HMI tags "Tabla de variables estándar_1"
   "MC066_STD" : , 1 s
   "MV031_STD" : , 1 s
   "MV032_STD" : , 1 s
   "MV030_STD" : , 1 s
   "DIP_1" : , internal
   "MP016_STD" : , 1 s
   "MC004_STD" : , 1 s
   "MP013_STD" : , 1 s
   "MV033_STD" : , 1 s
   "MC001_STD" : , 1 s
   "MC060_STD" : , 1 s
   "MC002_STD" : , 1 s
   "MP012_STD" : , 1 s
   "MC065_STD" : , 1 s
   "MS051_STD" : , 1 s
   "MC006_STD" : , 1 s
   "MP011_STD" : , 1 s
   "Iluminati_STD" : , 1 s
   "MC064_STD" : , 1 s
   "MS052_STD" : , 1 s
   "MT010_STD" : , 1 s
   "MS053_STD" : , 1 s
   "MP019_STD" : , 1 s
   "MC005_STD" : , 1 s
   "MC061_STD" : , 1 s
   "MV034_STD" : , 1 s
   "MC063_STD" : , 1 s
   "MP015_STD" : , 1 s
   "MT007_STD" : , 1 s
   "MS055_STD" : , 1 s
   "MP018_STD" : , 1 s
   "MP014_STD" : , 1 s
   "MS054_STD" : , 1 s
   "MS050_STD" : , 1 s
   "MP010_STD" : , 1 s
   "MT008_STD" : , 1 s
   "MT009_STD" : , 1 s
   "MC003_STD" : , 1 s
   "MC062_STD" : , 1 s
   "EB5" : Word, 1 s
   "EB7" : Word, 1 s
   "EB4" : Word, 1 s
   "EW8" : Word, 1 s
   "ACK_ALARMA_2" : Int, 1 s
   "MP020_STD" : Word, 1 s
   "MP021_STD" : Word, 1 s
   "MP022_STD" : Word, 1 s
   "CERO" : Bool, 1 s
   "UNO" : Bool, 1 s
   "IndCh" : Bool, 1 s
   "IndTrCh" : Bool, 1 s
   "IndCmpBaja" : Bool, 1 s
   "IndSecBaja" : Bool, 1 s
   "IndCmpAlta" : Bool, 1 s
   "IndSecAlta" : Bool, 1 s
   "IndTrCav" : Bool, 1 s
   "AnularSirena?" : Bool, internal
   "HorasBoost1" : DInt, 1 s
   "HorasBoost2" : DInt, 1 s
   "BoostPrHoras" : Bool, 1 s
   "BoostInvP" : Bool, 1 s
   "PrioridadBoost1" : Int, 1 s
   "PrioridadBoost2" : Int, 1 s
   "BoostInvPMan" : Bool, 1 s
   "min_boost1" : Int, 1 s
   "SegsBoost1" : Int, 1 s
   "SegsBoost" : Int, 1 s
   "MinBoost2" : Int, 1 s
   "FT1_AGUA" : Bool = PLC "FT1_AGUA", 1 s

HMI tags "AlarmasMTA"
   "AlarmasWord0" : Int, 1 s
   "AlarmasWord1" : Int, 1 s
   "AlarmasWord2" : Int, 1 s
   "AlarmasWord3" : Int, 1 s
   "AlarmasWord4" : Int, 1 s
   "AlarmasWord5" : Int, 1 s
   "AlarmasWord6" : Int, 1 s
   "AlarmasWord7" : Int, 1 s
   "AlarmasWord8" : Int, 1 s
   "Rec0" : Int, 1 s
   "Rec1" : Int, 1 s
   "Rec2" : Int, 1 s
   "Rec3" : Int, 1 s
   "Rec4" : Int, 1 s
   "Rec5" : Int, 1 s
   "Rec6" : Int, 1 s
   "Rec7" : Int, 1 s
   "Rec8" : Int, 1 s
   "AlarmasWord9" : Int, 1 s
   "AlarmasWord10" : Int, 1 s
   "AlarmasWord11" : Int, 1 s
   "AlarmasWord12" : Int, 1 s
   "AlarmasWord13" : Int, 1 s
   "AlarmasWord14" : Int, 1 s
   "Rec9" : Int, 1 s
   "Rec10" : Int, 1 s
   "Rec11" : Int, 1 s
   "Rec12" : Int, 1 s
   "Rec13" : Int, 1 s
   "Rec14" : Int, 1 s
   "AlarmasWord15" : Int, 1 s
   "Rec15" : Int, 1 s
   "ReconocerTODAS" : Bool, 1 s
   "EncendidoPLC" : Bool, 1 s
   "AlarmasWord16" : Int, 1 s
   "Rec16" : Int, 1 s
   "ReconocerTODAS_1" : Bool, 1 s
   "AlarmasWord18" : Int, 1 s
   "Rec18" : Int, 1 s
   "AlarmasWord19" : Int, 1 s
   "Rec19" : Int, 1 s
   "AlarmasWord20" : Int, 1 s
   "AlarmasWord21" : Int, 1 s
   "AlarmasWord22" : Int, 1 s
   "AlarmasWord23" : Int, 1 s
   "AlarmasWord24" : Int, 1 s
   "Rec20" : Int, 1 s
   "Rec21" : Int, 1 s
   "Rec22" : Int, 1 s
   "Rec23" : Int, 1 s
   "Rec24" : Int, 1 s

HMI tags "AutoTorresCav"
   "AutoV030" : Bool, 1 s
   "AutoV031" : Bool, 1 s
   "SP-OFF-V030" : Int, 1 s
   "SP-OFF-V031" : Int, 1 s
   "SP-ON-V030" : Int, 1 s
   "SP-ON-V031" : Int, 1 s

HMI tags "AutoTorresChillers"
   "AutoV001" : Bool, 1 s
   "AutoV002" : Bool, 1 s
   "AutoV003" : Bool, 1 s
   "SP-ON-V001" : Int, 1 s
   "SP-ON-V002" : Int, 1 s
   "SP-ON-V003" : Int, 1 s
   "SP-OFF-V001" : Int, 1 s
   "SP-OFF-V002" : Int, 1 s
   "SP-OFF-V003" : Int, 1 s
   "TemperaturatorresCH" : Real, 1 s

HMI tags "Booster"
   "AlarmaBooster" : Bool, 1 s
   "Booster_ModoManten" : Bool, 1 s
   "Booster_ModoManual" : Bool, 1 s
   "Booster_ModoAutoma" : Bool, 1 s
   "Booster_PlsManten" : Bool, 1 s
   "Booster_PlsManual" : Bool, 1 s
   "Booster_PlsAutoma" : Bool, 1 s
   "AnimaMotBooster" : Byte, 1 s
   "BoosterOrdMarcha" : Bool, 1 s
   "Booster_Conf_Marcha" : Bool, 1 s
   "Booster_Presost_Ctrl" : Bool, 1 s
   "Booster_Presost_PA" : Bool, 1 s
   "Booster_Habilitacion" : Bool, 1 s
   "Booster2_Conf_Marcha" : Bool, 1 s
   "Booster2_Habilitacion" : Bool, 1 s
   "Booster2_ModoAutoma" : Bool, 1 s
   "Booster2_ModoManten" : Bool, 1 s
   "Booster2_ModoManual" : Bool, 1 s
   "Booster2_PlsAutoma" : Bool, 1 s
   "Booster2_PlsManten" : Bool, 1 s
   "Booster2_PlsManual" : Bool, 1 s
   "AnimaMotBooster2" : Byte, 1 s
   "Booster2OrdMarcha" : Bool, 1 s
   "TiempoAyudaON" : Int, 1 s
   "TiempoAyudaOFF" : Int, 1 s
   "DifHorINVBoost" : DInt, 1 s
   "LimArrBoostPrio2" : Real, 1 s
   "LimArrBoostPrio1" : Real, 1 s
   "LimParBoostPrio2" : Real, 1 s
   "LimParBoostPrio1" : Real, 1 s
   "Presión_Actual_Boosters" : Real, 1 s
   "Ctrl_Analógico" : Bool, 1 s
   "Ver_Config" : Bool, internal
   "CotaSupPresAna" : Real, 1 s

HMI tags "CFG-Analog-MTA"
   "PresiónALTA" : Real, 1 s
   "PresiónBAJA" : Real, 1 s
   "TempCAV" : Real, 1 s
   "TempCH" : Real, 1 s
   "CFG-ALtaHH" : Real, 1 s
   "CFG-ALtaH" : Real, 1 s
   "CFG-ALtaL" : Real, 1 s
   "CFG-ALtaLL" : Real, 1 s
   "CFG-BajaHH" : Real, 1 s
   "CFG-BajaH" : Real, 1 s
   "CFG-BajaL" : Real, 1 s
   "CFG-BajaLL" : Real, 1 s
   "LO_potencia" : Real, 1 s
   "HI_caudal" : Real, 1 s
   "LO_caudal" : Real, 1 s
   "HI_potencia" : Real, 1 s
   "Caudal" : Real, 1 s
   "Potencia" : Real, 1 s

HMI tags "ChillersMTA"
   "HabMT007" : Bool, 1 s
   "HabMT008" : Bool, 1 s
   "HabMT009" : Bool, 1 s
   "HabMT010" : Bool, 1 s
   "DesMT007" : Bool, 1 s
   "DesMT008" : Bool, 1 s
   "DesMT009" : Bool, 1 s
   "DesMT010" : Bool, 1 s
   "MarchaMT007" : Bool, 1 s
   "MarchaMT008" : Bool, 1 s
   "MarchaMT009" : Bool, 1 s
   "MarchaMT010" : Bool, 1 s
   "ParadaMT007" : Bool, 1 s
   "ParadaMT008" : Bool, 1 s
   "ParadaMT009" : Bool, 1 s
   "ParadaMT010" : Bool, 1 s
   "Habilitación-CH-SOP-GR" : Bool, 1 s
   "Habilitación-CH-SOP-CH" : Bool, 1 s
   "Habilitación-CH-ENV-GR" : Bool, 1 s
   "Habilitación-CH-ENV-CH" : Bool, 1 s
   "Alarma1-CH-SOP-GR" : Bool, 1 s
   "Alarma2-CH-SOP-GR" : Bool, 1 s
   "RUN-CH-SOP-GR" : Bool, 1 s
   "MAX-CH-SOP-GR" : Bool, 1 s
   "AnimaciónMT007" : Byte, 1 s
   "AnimaciónMT008" : Byte, 1 s
   "AnimaciónMT009" : Byte, 1 s
   "AnimaciónMT010" : Byte, 1 s
   "AnimaciónMP010" : Byte, 1 s
   "AnimaciónMP011" : Byte, 1 s
   "AnimaciónMP012" : Byte, 1 s
   "AnimaciónMP013" : Byte, 1 s
   "HabMP010" : Bool, 1 s
   "HabMP011" : Bool, 1 s
   "HabMP012" : Bool, 1 s
   "HabMP013" : Bool, 1 s
   "HabMP018" : Bool, 1 s
   "HabMP019" : Bool, 1 s
   "DesMP010" : Bool, 1 s
   "DesMP011" : Bool, 1 s
   "DesMP012" : Bool, 1 s
   "DesMP013" : Bool, 1 s
   "DesMP018" : Bool, 1 s
   "DesMP019" : Bool, 1 s
   "MarchaMP010" : Bool, 1 s
   "MarchaMP011" : Bool, 1 s
   "MarchaMP012" : Bool, 1 s
   "MarchaMP013" : Bool, 1 s
   "MarchaMP018" : Bool, 1 s
   "MarchaMP019" : Bool, 1 s
   "ParadaMP010" : Bool, 1 s
   "ParadaMP011" : Bool, 1 s
   "ParadaMP012" : Bool, 1 s
   "ParadaMP013" : Bool, 1 s
   "ParadaMP018" : Bool, 1 s
   "ParadaMP019" : Bool, 1 s
   "AnimaciónMP018" : Byte, 1 s
   "AnimaciónMP019" : Byte, 1 s
   "DesV001" : Bool, 1 s
   "DesV002" : Bool, 1 s
   "HabV001" : Bool, 1 s
   "HabV002" : Bool, 1 s
   "MarchaV001" : Bool, 1 s
   "MarchaV002" : Bool, 1 s
   "ParadaV001" : Bool, 1 s
   "ParadaV002" : Bool, 1 s
   "AnimaciónV001" : Byte, 1 s
   "AnimaciónV002" : Byte, 1 s
   "VentiladoresMTA" : Bool, internal
   "MAX-CH-ENV-GR" : Bool, 1 s
   "RUN-CH-ENV-GR" : Bool, 1 s
   "Alarma2-CH-ENV-GR" : Bool, 1 s
   "Alarma1-CH-ENV-GR" : Bool, 1 s
   "SirenaM1" : Bool, 1 s
   "SirenaM2" : Bool, 1 s
   "SirenaM3" : Bool, 1 s
   "SirenaM4" : Bool, 1 s
   "AnimaciónV003" : Byte, 1 s
   "HabV003" : Bool, 1 s
   "DesV003" : Bool, 1 s
   "MarchaV003" : Bool, 1 s
   "ParadaV003" : Bool, 1 s
   "BombaTorreON" : Bool, 1 s
   "SirenaM5" : Bool, 1 s
   "SirenaChillers" : Bool, 1 s
   "SirenaM6" : Bool, 1 s
   "SirenaM7" : Bool, 1 s
   "SirenaM8" : Bool, 1 s
   "SirenaM9" : Bool, 1 s
   "SirenaM10" : Bool, 1 s
   "AlarmaNueva" : Bool, 1 s
   "AlarmaPresente" : Bool, 1 s
   "SinAlarmas" : Bool, 1 s
   "AlarmaAceite-CH-ENV-CH" : Bool, 1 s
   "AlarmaTemp-CH-ENV-CH" : Bool, 1 s
   "RUN-CH-ENV-CH" : Bool, 1 s
   "VerCh1MTA" : Bool, internal
   "VerCh2MTA" : Bool, internal
   "VerCh3MTA" : Bool, internal
   "VerCh4MTA" : Bool, internal
   "AlarmaPRUEBA" : DWord, 1 s
   "Presosato" : Bool, 1 s
   "CH-SOP-CH-CTC1ON" : Bool, 1 s
   "CH-SOP-CH-CTC2ON" : Bool, 1 s
   "CH-SOP-CH-TERM1" : Bool, 1 s
   "CH-SOP-CH-TERM2" : Bool, 1 s
   "CH-ENV-CH-ACT" : Bool, 1 s
   "CH-ENV-CH-TEMP" : Bool, 1 s
   "CH-ENV-CH-TERM" : Bool, 1 s
   "CH-ENV-CH-RUN" : Bool, 1 s
   "BombaTorreON2" : Bool, 1 s
   "HabV001(1)" : Bool, 1 s
   "HabV002(1)" : Bool, 1 s
   "HabV003(1)" : Bool, 1 s
   "HabV4" : Bool, 1 s
   "MarchaV001(1)" : Bool, 1 s
   "MarchaV002(1)" : Bool, 1 s
   "MarchaV003(1)" : Bool, 1 s
   "ParadaV001(1)" : Bool, 1 s
   "ParadaV002(1)" : Bool, 1 s
   "ParadaV003(1)" : Bool, 1 s
   "AnimaMenuV001" : Int, 1 s
   "AnimaMenuV002" : Int, 1 s
   "AnimaMenuV003" : Int, 1 s
   "DeshV001" : Bool, 1 s
   "DeshV002" : Bool, 1 s
   "DeshV003" : Bool, 1 s

HMI tags "CompBajaMTA"
   "HabilitaciónMC060" : Bool, 1 s
   "HabilitaciónMC061" : Bool, 1 s
   "HabilitaciónMC062" : Bool, 1 s
   "HabilitaciónMC063" : Bool, 1 s
   "HabilitaciónMC064" : Bool, 1 s
   "HabilitaciónMC065" : Bool, 1 s
   "DeshabilitaciónMC060" : Bool, 1 s
   "DeshabilitaciónMC061" : Bool, 1 s
   "DeshabilitaciónMC062" : Bool, 1 s
   "DeshabilitaciónMC063" : Bool, 1 s
   "DeshabilitaciónMC064" : Bool, 1 s
   "DeshabilitaciónMC065" : Bool, 1 s
   "MarchaMC060" : Bool, 1 s
   "MarchaMC061" : Bool, 1 s
   "MarchaMC062" : Bool, 1 s
   "MarchaMC063" : Bool, 1 s
   "MarchaMC064" : Bool, 1 s
   "MarchaMC065" : Bool, 1 s
   "ParadaMC060" : Bool, 1 s
   "ParadaMC061" : Bool, 1 s
   "ParadaMC062" : Bool, 1 s
   "ParadaMC063" : Bool, 1 s
   "ParadaMC064" : Bool, 1 s
   "ParadaMC065" : Bool, 1 s
   "AnimaMC060" : Byte, 1 s
   "AnimaMC061" : Byte, 1 s
   "AnimaMC062" : Byte, 1 s
   "AnimaMC063" : Byte, 1 s
   "AnimaMC064" : Byte, 1 s
   "AnimaMC065" : Byte, 1 s
   "VerMC060" : Bool, internal
   "VerMC061" : Bool, internal
   "VerMC062" : Bool, internal
   "VerMC063" : Bool, internal
   "VerMC064" : Bool, internal
   "MantM060" : Bool, 1 s
   "MantM061" : Bool, 1 s
   "MantM062" : Bool, 1 s
   "MantM063" : Bool, 1 s
   "MantM064" : Bool, 1 s
   "AutoMC060" : Bool, 1 s
   "AutoMC061" : Bool, 1 s
   "AutoMC062" : Bool, 1 s
   "AutoMC063" : Bool, 1 s
   "AutoMC064" : Bool, 1 s
   "SponMC060" : Real, 1 s
   "SponMC061" : Real, 1 s
   "SponMC062" : Real, 1 s
   "SponMC063" : Real, 1 s
   "SponMC064" : Real, 1 s
   "SpoffMC060" : Real, 1 s
   "SpoffMC061" : Real, 1 s
   "SpoffMC062" : Real, 1 s
   "SpoffMC063" : Real, 1 s
   "SpoffMC064" : Real, 1 s
   "AnimMenuMC060" : Int, 1 s
   "AnimMenuMC061" : Int, 1 s
   "AnimMenuMC062" : Int, 1 s
   "AnimMenuMC063" : Int, 1 s
   "AnimMenuMC064" : Int, 1 s
   "HabilitarMC060" : Bool, 1 s
   "AnularSirenaCav" : Bool, 1 s
   "VerMC65" : Bool, internal

HMI tags "CompresoresAltaMTA"
   "Sop1" : Bool, 1 s
   "Sop2" : Bool, 1 s
   "Sop3" : Bool, 1 s
   "ReqSop1" : Int, 1 s
   "ReqSop2" : Int, 1 s
   "ReqSop3" : Int, 1 s
   "NinSop" : Bool, 1 s
   "VCMP1" : Int, 1 s
   "VCMP2" : Int, 1 s
   "VCMP3" : Int, 1 s
   "VCMP4" : Int, 1 s
   "VCMP5" : Int, 1 s
   "IncP1" : Bool, 100 ms
   "IncP2" : Bool, 100 ms
   "IncP3" : Bool, 100 ms
   "IncP4" : Bool, 100 ms
   "IncP5" : Bool, 100 ms
   "DecP1" : Bool, 1 s
   "DecP2" : Bool, 1 s
   "DecP3" : Bool, 1 s
   "DecP4" : Bool, 1 s
   "DecP5" : Bool, 1 s
   "PriRealCMP1" : Int, 1 s
   "PriRealCMP2" : Int, 1 s
   "PriRealCMP3" : Int, 1 s
   "PriRealCMP4" : Int, 1 s
   "PriRealCMP5" : Int, 1 s
   "Auto1" : Bool, 1 s
   "Auto2" : Bool, 1 s
   "Auto3" : Bool, 1 s
   "Auto4" : Bool, 1 s
   "Auto5" : Bool, 1 s
   "IndV1" : Bool, 100 ms
   "IndV2" : Bool, 100 ms
   "IndV3" : Bool, 100 ms
   "IndV4" : Bool, 100 ms
   "IndV5" : Bool, 100 ms
   "IndR1" : Bool, 100 ms
   "IndR2" : Bool, 100 ms
   "IndR3" : Bool, 100 ms
   "IndR4" : Bool, 100 ms
   "IndR5" : Bool, 100 ms
   "Est1" : Word, 1 s
   "Est2" : Word, 1 s
   "Est3" : Word, 1 s
   "Est4" : Word, 1 s
   "Est5" : Word, 1 s
   "LimSUP1" : Real, 1 s
   "LimSUP2" : Real, 1 s
   "LimSUP3" : Real, 1 s
   "LimSUP4" : Real, 1 s
   "LimSUP5" : Real, 1 s
   "LimINF1" : Real, 1 s
   "LimINF2" : Real, 1 s
   "LimINF3" : Real, 1 s
   "LimINF4" : Real, 1 s
   "LimINF5" : Real, 1 s
   "PresMaX" : Real, 1 s
   "Delta" : Real, 1 s
   "Hist" : Real, 1 s
   "CompReq" : Int, 1 s
   "CompReqINI" : Int, 1 s
   "AnimMenuMC001" : Int, 1 s
   "AnimMenuMC002" : Int, 1 s
   "AnimMenuMC003" : Int, 1 s
   "AnimMenuMC004" : Int, 1 s
   "AnimMenuMC005" : Int, 1 s
   "SPON1" : Real, 1 s
   "SPON2" : Real, 1 s
   "SPON3" : Real, 1 s
   "SPON4" : Real, 1 s
   "SPON5" : Real, 1 s
   "SPOFF1" : Real, 1 s
   "SPOFF2" : Real, 1 s
   "SPOFF3" : Real, 1 s
   "SPOFF4" : Real, 1 s
   "SPOFF5" : Real, 1 s
   "MantMC001" : Bool, 1 s
   "MantMC002" : Bool, 1 s
   "MantMC003" : Bool, 1 s
   "MantMC004" : Bool, 1 s
   "MantMC005" : Bool, 1 s
   "IndVparp1" : Bool, 1 s
   "IndVparp2" : Bool, 1 s
   "IndVparp3" : Bool, 1 s
   "IndVparp4" : Bool, 1 s
   "IndVparp5" : Bool, 1 s
   "TiempoenVacío" : Int, 1 s
   "TiemposinReq" : Int, 1 s
   "TiempoSop" : Int, 1 s
   "HistCRT" : Real, 1 s
   "LimINFCRT" : Real, 1 s
   "LimSUPCRT" : Real, 1 s
   "PanMCH1" : Bool, 1 s
   "PanMCH2" : Bool, 1 s
   "PanMCH3" : Bool, 1 s
   "PanMCH4" : Bool, 1 s
   "PanMCH5" : Bool, 1 s
   "MarchaMC001" : Bool, 1 s
   "MarchaMC002" : Bool, 1 s
   "MarchaMC003" : Bool, 1 s
   "MarchaMC004" : Bool, 1 s
   "MarchaMC005" : Bool, 1 s
   "ParadaMC001" : Bool, 1 s
   "ParadaMC002" : Bool, 1 s
   "ParadaMC003" : Bool, 1 s
   "ParadaMC004" : Bool, 1 s
   "ParadaMC005" : Bool, 1 s
   "AnimMotorMC001" : Byte, 1 s
   "AnimMotorMC002" : Byte, 1 s
   "AnimMotorMC003" : Byte, 1 s
   "AnimMotorMC004" : Byte, 1 s
   "AnimMotorMC005" : Byte, 1 s
   "EV1" : Bool, 1 s
   "EV2" : Bool, 1 s
   "EV3" : Bool, 1 s
   "EV4" : Bool, 1 s
   "EV5" : Bool, 1 s
   "HORAS1" : DInt, 1 s
   "HORAS2" : DInt, 1 s
   "HORAS3" : DInt, 1 s
   "HORAS4" : DInt, 1 s
   "HORAS5" : DInt, 1 s
   "MIN1" : Int, 1 s
   "MIN2" : Int, 1 s
   "MIN3" : Int, 1 s
   "MIN4" : Int, 1 s
   "MIN5" : Int, 1 s
   "MarchaOK1" : Bool, 1 s
   "MarchaOK2" : Bool, 1 s
   "MarchaOK3" : Bool, 1 s
   "MarchaOK4" : Bool, 1 s
   "MarchaOK5" : Bool, 1 s
   "ForzarMarcha1" : Bool, 1 s
   "ForzarMarcha2" : Bool, 1 s
   "ForzarMarcha3" : Bool, 1 s
   "ForzarMarcha4" : Bool, 1 s
   "ForzarMarcha5" : Bool, 1 s
   "ForzarParada1" : Bool, 1 s
   "ForzarParada2" : Bool, 1 s
   "ForzarParada3" : Bool, 1 s
   "ForzarParada4" : Bool, 1 s
   "ForzarParada5" : Bool, 1 s
   "SPONF1" : Real, 1 s
   "SPONF2" : Real, 1 s
   "SPONF3" : Real, 1 s
   "SPONF4" : Real, 1 s
   "SPONF5" : Real, 1 s
   "SPOFFF1" : Real, 1 s
   "SPOFFF2" : Real, 1 s
   "SPOFFF3" : Real, 1 s
   "SPOFFF4" : Real, 1 s
   "SPOFFF5" : Real, 1 s
   "ForzandoMarcha1" : Bool, 1 s
   "ForzandoMarcha2" : Bool, 1 s
   "ForzandoMarcha3" : Bool, 1 s
   "ForzandoMarcha4" : Bool, 1 s
   "ForzandoMarcha5" : Bool, 1 s
   "MediaCargaBellis" : Bool, 1 s
   "SPONF3b" : Real, 1 s
   "SPOFFF3b" : Real, 1 s
   "EV3b" : Bool, 1 s
   "TiempoMaxBellismedia" : Int, 1 s
   "Est6" : Int, 1 s
   "PriRealCMP6" : Int, 1 s
   "IndV6" : Bool, 1 s

HMI tags "IluminaciónMTA"
   "TiempoIluminación" : Word, 1 s
   "EncendidoPanel" : Bool, 1 s
   "ApagadoPanel" : Bool, 1 s
   "ON" : Bool, 1 s
   "MantenerON" : Bool, 1 s
   "AlarmaBoosters" : Bool, 1 s

HMI tags "SecadoresAltaMTA"
   "AnimaMS050" : Byte, 1 s
   "AnimaMS051" : Byte, 1 s
   "AnimaMS052" : Byte, 1 s
   "AnimaMS053" : Byte, 1 s
   "DeshabilitaciónMS050" : Bool, 1 s
   "DeshabilitaciónMS051" : Bool, 1 s
   "DeshabilitaciónMS052" : Bool, 1 s
   "DeshabilitaciónMS053" : Bool, 1 s
   "HabilitaciónMS050" : Bool, 1 s
   "HabilitaciónMS051" : Bool, 1 s
   "HabilitaciónMS052" : Bool, 1 s
   "HabilitaciónMS053" : Bool, 1 s
   "MantMS050" : Bool, 1 s
   "MantMS051" : Bool, 1 s
   "MantMS052" : Bool, 1 s
   "MantMS053" : Bool, 1 s
   "MarchaMS050" : Bool, 1 s
   "MarchaMS051" : Bool, 1 s
   "MarchaMS052" : Bool, 1 s
   "MarchaMS053" : Bool, 1 s
   "ParadaMS050" : Bool, 1 s
   "ParadaMS051" : Bool, 1 s
   "ParadaMS052" : Bool, 1 s
   "ParadaMS053" : Bool, 1 s
   "AnimaMenuMS050" : Int, 1 s
   "AnimaMenuMS051" : Int, 1 s
   "AnimaMenuMS052" : Int, 1 s
   "AnimaMenuMS053" : Int, 1 s
   "Enc1MS050" : Int, 1 s
   "Enc2MS050" : Int, 1 s
   "Enc1MS051" : Int, 1 s
   "Enc2MS051" : Int, 1 s
   "Enc1MS052" : Int, 1 s
   "Enc2MS052" : Int, 1 s
   "Enc1MS053" : Int, 1 s
   "Enc2MS053" : Int, 1 s
   "AutoMS050" : Bool, 1 s
   "AutoMS051" : Bool, 1 s
   "AutoMS052" : Bool, 1 s
   "AutoMS053" : Bool, 1 s

HMI tags "SecadoresBaja"
   "AnimaMS054" : Byte, 1 s
   "AnimaMS055" : Byte, 1 s
   "DeshabilitaciónMS054" : Bool, 1 s
   "DeshabilitaciónMS055" : Bool, 1 s
   "HabilitaciónMS054" : Bool, 1 s
   "HabilitaciónMS055" : Bool, 1 s
   "MarchaMS054" : Bool, 1 s
   "MarchaMS055" : Bool, 1 s
   "ParadaMS054" : Bool, 1 s
   "ParadaMS055" : Bool, 1 s
   "MantMS054" : Bool, 1 s
   "MantMS055" : Bool, 1 s

HMI tags "SENTRON PAC 3200"
   "Tension Fase R" : Float, 1 s
   "Tension fase S" : Float, 1 s
   "Tension Fase T" : Float, 1 s
   "Tension Linea RS" : Float, 1 s
   "Tension Linea ST" : Float, 1 s
   "Tension Linea TR" : Float, 1 s
   "Corriente fase R" : Float, 1 s
   "Corriente Fase S" : Float, 1 s
   "Corriente Fase T" : Float, 1 s
   "Pot.Apa R" : Float, 1 s
   "Pot.Apa S" : Float, 1 s
   "Pot.Apa T" : Float, 1 s
   "Pot.Act R" : Float, 1 s
   "Pot.Act S" : Float, 1 s
   "Pot.Act T" : Float, 1 s
   "Pot.ReAct R" : Float, 1 s
   "Pot.ReAct S" : Float, 1 s
   "Pot.ReAct T" : Float, 1 s
   "Coseno R" : Float, 1 s
   "Coseno S" : Float, 1 s
   "Coseno T" : Float, 1 s
   "THD-R TensionFase R" : Float, 1 s
   "THD-R Tension Fase S" : Float, 1 s
   "THD-R Tension Fase T" : Float, 1 s
   "THD-R Corriente Fase R" : Float, 1 s
   "THD-R Corriente Fase S" : Float, 1 s
   "THD-R Corriente Fase T" : Float, 1 s
   "Frecuencia" : Float, 1 s
   "Tension Media Fase" : Float, 1 s
   "Tension Media de Linea" : Float, 1 s
   "Corriente Media" : Float, 1 s
   "Pot Apa Total" : Float, 1 s
   "Pot Act Total" : Float, 1 s
   "Pot ReAct Total" : Float, 1 s
   "coseno Total" : Float, 1 s
   "desbalance de tension" : Float, 1 s
   "desbalance de corriente" : Float, 1 s
   "Tension Maxima R" : Float, 1 s
   "Tension Maxima S" : Float, 1 s
   "Tension Maxima T" : Float, 1 s
   "Tension Maxima RS" : Float, 1 s
   "Tension Maxima ST" : Float, 1 s
   "Tension Maxima TR" : Float, 1 s
   "Corriente Maxima R" : Float, 1 s
   "Corriente Maxima S" : Float, 1 s
   "Corriente Maxima T" : Float, 1 s

HMI tags "TorresCav-MTA"
   "AnimaMV030" : Byte, 1 s
   "AnimaMV031" : Byte, 1 s
   "AnimaMP014" : Byte, 1 s
   "AnimaMP015" : Byte, 1 s
   "DeshabilitaciónMV030" : Bool, 1 s
   "DeshabilitaciónMV031" : Bool, 1 s
   "DeshabilitaciónMP014" : Bool, 1 s
   "DeshabilitaciónMP015" : Bool, 1 s
   "HabilitaciónMV030" : Bool, 1 s
   "HabilitaciónMV031" : Bool, 1 s
   "HabilitaciónMP014" : Bool, 1 s
   "HabilitaciónMP015" : Bool, 1 s
   "MantMV030" : Bool, 1 s
   "MantMV031" : Bool, 1 s
   "MantMP014" : Bool, 1 s
   "MantMP015" : Bool, 1 s
   "MarchaMV030" : Bool, 1 s
   "MarchaMV031" : Bool, 1 s
   "MarchaMP014" : Bool, 1 s
   "MarchaMP015" : Bool, 1 s
   "ParadaMV030" : Bool, 1 s
   "ParadaMV031" : Bool, 1 s
   "ParadaMP014" : Bool, 1 s
   "ParadaMP015" : Bool, 1 s
   "MenuV030" : Int, 1 s
   "MenuV031" : Int, 1 s

discrete alarms
   1: '', class MTA, trigger "AlarmasWord13" bit 9
   2: '', class MTA, trigger "AlarmasWord13" bit 10
   3: '', class MTA, trigger "AlarmasWord13" bit 11
   4: '', class MTA, trigger "AlarmasWord13" bit 12
   5: '', class MTA, trigger "AlarmasWord13" bit 13
   6: '', class MTA, trigger "AlarmasWord13" bit 14
   7: '', class MTA, trigger "AlarmasWord13" bit 15
   8: '', class MTA, trigger "AlarmasWord14" bit 8
   9: '', class MTA, trigger "AlarmasWord14" bit 9
   10: '', class MTA, trigger "AlarmasWord14" bit 10
   11: '', class MTA, trigger "AlarmasWord14" bit 11
   12: '', class MTA, trigger "AlarmasWord14" bit 12
   13: '', class MTA, trigger "AlarmasWord6" bit 8
   14: '', class MTA, trigger "AlarmasWord6" bit 9
   15: '', class MTA, trigger "AlarmasWord14" bit 13
   16: '', class MTA, trigger "AlarmasWord14" bit 14
   17: '', class MTA, trigger "AlarmasWord14" bit 15
   18: '', class MTA, trigger "AlarmasWord15" bit 8
   19: '', class MTA, trigger "AlarmasWord15" bit 9
   20: '', class MTA, trigger "AlarmasWord15" bit 10
   21: '', class MTA, trigger "AlarmasWord15" bit 11
   22: '', class MTA, trigger "AlarmasWord15" bit 12
   23: '', class MTA, trigger "AlarmasWord15" bit 13
   24: '', class MTA, trigger "AlarmasWord15" bit 14
   25: '', class MTA, trigger "AlarmasWord15" bit 15
   26: '', class MTA, trigger "AlarmasWord16" bit 8
   27: '', class MTA, trigger "AlarmasWord16" bit 9
   28: '', class MTA, trigger "AlarmasWord16" bit 10
   29: '', class MTA, trigger "AlarmasWord16" bit 11
   30: '', class MTA, trigger "AlarmasWord16" bit 12
   31: '', class MTA, trigger "AlarmasWord16" bit 13
   32: '', class MTA, trigger "AlarmasWord16" bit 14
   33: '', class MTA, trigger "AlarmasWord16" bit 15
   50: '', class MTA, trigger "AlarmasWord6" bit 10
   53: '', class MTA, trigger "AlarmasWord6" bit 11
   66: '', class MTA, trigger "AlarmasWord7" bit 8
   67: '', class MTA, trigger "AlarmasWord7" bit 9
   68: '', class MTA, trigger "AlarmasWord7" bit 10
   69: '', class MTA, trigger "AlarmasWord7" bit 11
   70: '', class MTA, trigger "AlarmasWord7" bit 12
   71: '', class MTA, trigger "AlarmasWord7" bit 13
   72: '', class MTA, trigger "AlarmasWord7" bit 14
   73: '', class MTA, trigger "AlarmasWord7" bit 15
   74: '', class MTA, trigger "AlarmasWord8" bit 8
   75: '', class MTA, trigger "AlarmasWord8" bit 9
   76: '', class MTA, trigger "AlarmasWord8" bit 10
   77: '', class MTA, trigger "AlarmasWord8" bit 11
   78: '', class MTA, trigger "AlarmasWord8" bit 12
   79: '', class MTA, trigger "AlarmasWord8" bit 13
   80: '', class MTA, trigger "AlarmasWord8" bit 14
   81: '', class MTA, trigger "AlarmasWord8" bit 15
   82: '', class MTA, trigger "AlarmasWord9" bit 8
   83: '', class MTA, trigger "AlarmasWord9" bit 9
   87: '', class MTA, trigger "AlarmasWord6" bit 12
   88: '', class MTA, trigger "AlarmasWord6" bit 13
   89: '', class MTA, trigger "AlarmasWord6" bit 14
   90: '', class MTA, trigger "AlarmasWord6" bit 15
   91: '', class MTA, trigger "AlarmasWord9" bit 10
   92: '', class MTA, trigger "AlarmasWord9" bit 11
   93: '', class MTA, trigger "AlarmasWord9" bit 12
   94: '', class MTA, trigger "AlarmasWord9" bit 13
   95: '', class MTA, trigger "AlarmasWord9" bit 14
   96: '', class MTA, trigger "AlarmasWord9" bit 15
   97: '', class MTA, trigger "AlarmasWord10" bit 8
   98: '', class MTA, trigger "AlarmasWord10" bit 9
   99: '', class MTA, trigger "AlarmasWord10" bit 10
   100: '', class MTA, trigger "AlarmasWord10" bit 11
   101: '', class MTA, trigger "AlarmasWord10" bit 12
   102: '', class MTA, trigger "AlarmasWord10" bit 13
   103: '', class MTA, trigger "AlarmasWord10" bit 14
   104: '', class MTA, trigger "AlarmasWord10" bit 15
   105: '', class MTA, trigger "AlarmasWord11" bit 8
   106: '', class MTA, trigger "AlarmasWord11" bit 9
   107: '', class MTA, trigger "AlarmasWord11" bit 10
   108: '', class MTA, trigger "AlarmasWord11" bit 11
   109: '', class MTA, trigger "AlarmasWord11" bit 12
   110: '', class MTA, trigger "AlarmasWord11" bit 13
   111: '', class MTA, trigger "AlarmasWord11" bit 14
   112: '', class MTA, trigger "AlarmasWord11" bit 15
   113: '', class MTA, trigger "AlarmasWord12" bit 8
   114: '', class MTA, trigger "AlarmasWord12" bit 9
   115: '', class MTA, trigger "AlarmasWord12" bit 10
   116: '', class MTA, trigger "AlarmasWord12" bit 11
   117: '', class MTA, trigger "AlarmasWord12" bit 12
   118: '', class MTA, trigger "AlarmasWord12" bit 13
   119: '', class MTA, trigger "AlarmasWord12" bit 14
   120: '', class MTA, trigger "AlarmasWord12" bit 15
   121: '', class MTA, trigger "AlarmasWord13" bit 8
   125: '', class MTA, trigger "AlarmasWord4" bit 8
   126: '', class MTA, trigger "AlarmasWord3" bit 15
   127: '', class MTA, trigger "AlarmasWord4" bit 11
   128: '', class MTA, trigger "AlarmasWord4" bit 10
   129: '', class MTA, trigger "AlarmasWord4" bit 9
   130: '', class MTA, trigger "AlarmasWord3" bit 11
   131: '', class MTA, trigger "AlarmasWord3" bit 10
   132: '', class MTA, trigger "AlarmasWord3" bit 9
   133: '', class MTA, trigger "AlarmasWord3" bit 14
   134: '', class MTA, trigger "AlarmasWord3" bit 13
   135: '', class MTA, trigger "AlarmasWord3" bit 12
   136: '', class MTA, trigger "AlarmasWord4" bit 12
   137: '', class MTA, trigger "AlarmasWord4" bit 15
   138: '', class MTA, trigger "AlarmasWord4" bit 14
   139: '', class MTA, trigger "AlarmasWord4" bit 13
   140: '', class MTA, trigger "AlarmasWord3" bit 8
   141: '', class MTA, trigger "AlarmasWord1" bit 8
   142: '', class MTA, trigger "AlarmasWord0" bit 15
   143: '', class MTA, trigger "AlarmasWord0" bit 14
   144: '', class MTA, trigger "AlarmasWord1" bit 11
   145: '', class MTA, trigger "AlarmasWord1" bit 10
   146: '', class MTA, trigger "AlarmasWord1" bit 9
   147: '', class MTA, trigger "AlarmasWord0" bit 10
   148: '', class MTA, trigger "AlarmasWord0" bit 9
   149: '', class MTA, trigger "AlarmasWord0" bit 8
   150: '', class MTA, trigger "AlarmasWord0" bit 13
   151: '', class MTA, trigger "AlarmasWord0" bit 12
   152: '', class MTA, trigger "AlarmasWord0" bit 11
   153: '', class MTA, trigger "AlarmasWord1" bit 12
   154: '', class MTA, trigger "AlarmasWord2" bit 12
   155: '', class MTA, trigger "AlarmasWord2" bit 11
   156: '', class MTA, trigger "AlarmasWord2" bit 10
   157: '', class MTA, trigger "AlarmasWord2" bit 15
   158: '', class MTA, trigger "AlarmasWord2" bit 14
   159: '', class MTA, trigger "AlarmasWord2" bit 13
   160: '', class MTA, trigger "AlarmasWord1" bit 15
   161: '', class MTA, trigger "AlarmasWord1" bit 14
   162: '', class MTA, trigger "AlarmasWord1" bit 13
   163: '', class MTA, trigger "AlarmasWord2" bit 9
   164: '', class MTA, trigger "AlarmasWord2" bit 8
   165: '', class MTA, trigger "AlarmasWord5" bit 8
   166: '', class MTA, trigger "AlarmasWord5" bit 9
   167: '', class MTA, trigger "AlarmasWord5" bit 10
   168: '', class MTA, trigger "AlarmasWord5" bit 11
   169: '', class MTA, trigger "AlarmasWord5" bit 12
   170: '', class MTA, trigger "AlarmasWord5" bit 13
   171: '', class MTA, trigger "AlarmasWord5" bit 14
   172: '', class MTA, trigger "AlarmasWord5" bit 15
   34: '', class MTA, trigger "AlarmasWord18" bit 8
   35: '', class MTA, trigger "AlarmasWord18" bit 9
   36: '', class MTA, trigger "AlarmasWord18" bit 10
   37: '', class MTA, trigger "AlarmasWord18" bit 11
   38: '', class MTA, trigger "AlarmasWord18" bit 12
   39: '', class MTA, trigger "AlarmasWord18" bit 13
   40: '', class MTA, trigger "AlarmasWord18" bit 14
   41: '', class MTA, trigger "Rec4" bit 15
   42: '', class MTA, trigger "AlarmasWord19" bit 8
   43: '', class MTA, trigger "AlarmasWord19" bit 9
   44: '', class MTA, trigger "AlarmasWord19" bit 10
   45: '', class MTA, trigger "AlarmasWord19" bit 11
   46: '', class MTA, trigger "AlarmasWord19" bit 12
   47: '', class MTA, trigger "AlarmasWord19" bit 13
   48: '', class MTA, trigger "AlarmasWord20" bit 8
   49: '', class MTA, trigger "AlarmasWord20" bit 9
   51: '', class MTA, trigger "AlarmasWord20" bit 10
   52: '', class MTA, trigger "AlarmasWord20" bit 11
   54: '', class MTA, trigger "AlarmasWord20" bit 12
   55: '', class MTA, trigger "AlarmasWord20" bit 13
   56: '', class MTA, trigger "AlarmasWord20" bit 14
   57: '', class MTA, trigger "AlarmasWord20" bit 15
   58: '', class MTA, trigger "AlarmasWord21" bit 8
   59: '', class MTA, trigger "AlarmasWord21" bit 9
   60: '', class MTA, trigger "AlarmasWord21" bit 10
   61: '', class MTA, trigger "AlarmasWord21" bit 11
   62: '', class MTA, trigger "AlarmasWord21" bit 12
   63: '', class MTA, trigger "AlarmasWord21" bit 13
   64: '', class MTA, trigger "AlarmasWord21" bit 14
   65: '', class MTA, trigger "AlarmasWord21" bit 15
   84: '', class MTA, trigger "AlarmasWord22" bit 8
   85: '', class MTA, trigger "AlarmasWord22" bit 9
   86: '', class MTA, trigger "AlarmasWord22" bit 10
   122: '', class MTA, trigger "AlarmasWord22" bit 11
   123: '', class MTA, trigger "AlarmasWord22" bit 12
   124: '', class MTA, trigger "AlarmasWord22" bit 13
   173: '', class MTA, trigger "AlarmasWord22" bit 14
   174: '', class MTA, trigger "AlarmasWord22" bit 15
   175: '', class MTA, trigger "AlarmasWord23" bit 8
   176: '', class MTA, trigger "AlarmasWord23" bit 9
   177: '', class MTA, trigger "AlarmasWord23" bit 10
   178: '', class MTA, trigger "AlarmasWord23" bit 11
   179: '', class MTA, trigger "AlarmasWord23" bit 12
   180: '', class MTA, trigger "AlarmasWord23" bit 13
   181: '', class MTA, trigger "AlarmasWord23" bit 14
   182: '', class MTA, trigger "AlarmasWord23" bit 15
   183: '', class MTA, trigger "AlarmasWord24" bit 8
   184: '', class MTA, trigger "AlarmasWord24" bit 9
   185: '', class MTA, trigger "AlarmasWord24" bit 10
   186: '', class MTA, trigger "AlarmasWord24" bit 11
   199: '', class MTA, trigger "AlarmasWord24" bit 15

text list "EstadoMotor": 0 ''; 1 ''; 2 ''; 3 ''; 4 ''; 5 ''; 6 ''; 7 ''

text list "EstadoCmpAlta": 256 ''; 512 ''; 1024 ''; 2048 ''; 4096 ''; 8192 ''; 16384 ''; 32768 ''; 1 ''

text list "Presostato Ctrl": 0 ''; 1 ''

text list "Presostato de Alarma": 0 ''; 1 ''

text list "Lista de rutas": 0 ''; 1 ''; 2 ''; 3 ''; 4 ''; 5 ''; 6 ''; 7 ''; 8 ''; 9 ''; 10 ''

text list "Lista de compresores": 0 ''; 1 ''; 2 ''; 3 ''; 4 ''; 5 ''; 6 ''; 7 ''; 8 ''; 9 ''; 10 ''

graphic list "Motor2": 0 'Motor2Dorado'; 1 'Motor2Verde_1'; 2 'Motor2VerdeOscuro'; 3 'Motor2Azul'; 4 'Motor2Celeste'; 5 'Motor2Amarillo'; 6 'Motor2Gris_1'; 7 'Motor2Rojo'; 8 'Motor2Dorado'

graphic list "MotorBelliss": 0 'dorado'; 1 'bell1ve'; 2 'bell1ve'; 3 'az'; 4 'az'; 5 'bell1am'; 6 'dorado'; 7 'az'

graphic list "BarraPrioridades": 1 'R1'; 2 'R2'; 3 'R3'; 4 'R4'; 5 'R5'; 6 'R4'; 6 'R6.rlu'

graphic list "Indicador": 0 'indDorado'; 1 'indVerde'; 2 'indVerde_1'; 3 'indAZUL'; 4 'indCeleste'; 5 'indAmarillo'; 6 'indGris'; 7 'indRojo'; 8 'indCeleste'

graphic list "BarraPrioridades_1": 1 'set1'; 2 'set2'; 3 'set3'; 4 'set4'; 5 'set5'; 6 'set4'; 6 'set6'

graphic list "BaseSullChico": 0 'BaseSullChicoDorado_4'; 1 'BaseSullChico'; 2 'BaseSullChico'; 3 'BaseSullChicoAzul_4'; 4 'BaseSullChicoAzul_4'; 5 'BaseSullChicoAmarillo_4'; 6 'BaseSullChicoGris_4'; 7 'BaseSullChicoRojo_4'; 8 'BaseSullChicoAzul_4'

graphic list "MotorTorre": 0 'torreFINAL4C2_1'; 1 'torreFINAL4C2v_2'; 2 'torreFINAL4C2v_2'; 3 'torreFINAL4C2b'; 4 'torreFINAL4C2b'; 5 'torreFINAL4C2a_2'; 6 'torreFINAL4C2_1'; 7 'torreFINAL4C2_1'

graphic list "Secador2": 0 'BaseSullChicoDorado_2'; 1 'BaseSullChico_5'; 2 'BaseSullChico_5'; 3 'BaseSullChicoAzul_2'; 4 'BaseSullChicoAzul_2'; 5 'BaseSullChicoAmarillo_2'; 6 'BaseSullChicoGris_2'; 7 'BaseSullChicoRojo_2'

graphic list "Secador1": 0 'BaseSullChicoDorado_1'; 1 'BaseSullChico_4'; 2 'BaseSullChico_4'; 3 'BaseSullChicoAzul_1'; 4 'BaseSullChicoAzul_1'; 5 'BaseSullChicoAmarillo_1'; 6 'BaseSullChicoGris_1'; 7 'BaseSullChicoRojo_1'

graphic list "Motor Grande": 0 'MotorDorado'; 1 'MotorVerde'; 2 'MotorVerde'; 3 'MotorAzul'; 4 'MotorCeleste'; 5 'MotorAmarillo'; 6 'MotorGris'; 7 'MotorRojo'; 8 'MotorCeleste'

graphic list "Mantenimiento": 0 'MECH2'; 1 'MECH1'

graphic list "Motor Chico": 0 'Booster-D-Dor2'; 1 'Booster-D-VE2'; 2 'Booster-D-VE2'; 3 'Booster-D-Azul2'; 4 'Booster-D-AZ2'; 5 'Booster-D-AM2'; 6 'Booster-D-GR'; 7 'Booster-D-RO2'; 8 'Booster-D-AZ2'

graphic list "Hélice": 0 'Booster-C1'; 1 'Booster-C2'

screen "Graf-Corrientes" 1280x800, template "Plantilla"
   TrendView "Visor de curvas_1" at 8,72 size 1260x636
   TextField "Campo de texto_16" at 493,10 size 294x27

screen "Graf-Fase" 1280x800, template "Plantilla"
   TrendView "Visor de curvas_1" at 3,65 size 1268x644
   TextField "Campo de texto_16" at 477,10 size 364x27

screen "Grafica" 1280x800, template "Plantilla"
   Button "Botón_7" at 368,280 size 240x49
   Button "Botón_12" at 367,440 size 240x49
   Button "Botón_13" at 368,216 size 240x49
   TextField "Campo de texto_1" at 55,108 size 353x27
   Button "Botón_1" at 767,280 size 240x49
   TextField "Campo de texto_16" at 521,10 size 226x27
   Button "Botón_2" at 368,344 size 240x49
   Button "Botón_3" at 766,440 size 240x49
   Button "Botón_4" at 769,526 size 240x49

screen "GraficaPALTA" 1280x800, template "Plantilla"
   TrendView "Visor de curvas_1" at 5,79 size 1234x618
   TextField "Campo de texto_16" at 521,10 size 193x27

screen "GraficaPBAJA" 1280x800, template "Plantilla"
   TrendView "Visor de curvas_1" at 5,71 size 1242x626
   TextField "Campo de texto_16" at 521,10 size 198x27

screen "GraficaTCAV" 1280x800, template "Plantilla"
   TrendView "Visor de curvas_1" at 5,71 size 1242x626
   TextField "Campo de texto_16" at 521,10 size 254x27

screen "GraficaTCH" 1280x800, template "Plantilla"
   TrendView "Visor de curvas_1" at 5,71 size 1242x626
   TextField "Campo de texto_16" at 521,10 size 243x27

screen "GraficaTodas" 1280x800, template "Plantilla"
   TrendView "Visor de curvas_1" at 5,71 size 1242x626

screen "Graf-Linea" 1280x800, template "Plantilla"
   TrendView "Visor de curvas_1" at 3,65 size 1268x652
   TextField "Campo de texto_16" at 453,10 size 370x27

screen "Graf-Pot" 1280x800, template "Plantilla"
   TrendView "Visor de curvas_1" at 3,65 size 1268x644
   TextField "Campo de texto_16" at 477,10 size 339x27

screen "Graf-PotTotal" 1280x800, template "Plantilla"
   TrendView "Visor de curvas_1" at 3,65 size 1268x644
   TextField "Campo de texto_16" at 477,10 size 327x27

screen "IluminaciónMTA" 1280x800, template "Plantilla"
   Switch "Interruptor_1" at 36,546 size 510x96
   Button "Botón_1" at 36,264 size 248x96
   Button "Botón_2" at 298,263 size 248x96
   IOField "Campo ES_1" at 257,148 size 140x39
   TextField "Campo de texto_1" at 42,156 size 186x27
   TextField "Campo de texto_3" at 58,190 size 466x58
   TextField "Campo de texto_2" at 58,414 size 433x112
   TextField "Campo de texto_16" at 553,10 size 177x27

screen "INICIO" 1280x800, template "Plantilla"
   Button "Botón_1" at 1025,513 size 108x65
   Button "Botón_2" at 115,501 size 130x47
   UserView "Visor de usuarios_1" at 266,510 size 665x23
   GraphicView "Visor de gráficos_1" at 96,110 size 1064x352
   Button "Botón_3" at 115,557 size 130x47
   Button "Botón_4" at 802,557 size 130x47

screen "INICIO-Administración" 1280x800, template "Plantilla"
   Button "Botón_1" at 1025,513 size 108x65
   Button "Botón_2" at 115,501 size 130x47
   UserView "Visor de usuarios_1" at 266,502 size 665x23
   GraphicView "Visor de gráficos_1" at 96,110 size 1064x352
   Button "Botón_3" at 115,557 size 130x47
   UserView "Visor de usuarios_2" at 266,534 size 665x143

screen "MTA-ALTAMC001" 1280x800, template "Plantilla-Alta-Cmp"
   Switch "Interruptor_1" at 156,166 size 37x37
   Button "Botón_6" at 27,153 size 88x62
   ScreenModuleView "Faceplate_6_1" at 348,235 size 76x34
   ScreenModuleView "Faceplate_7_1" at 208,157 size 216x70
   GraphicIOField "Campo ES gráfico_2" at 16,279 size 422x6
   SymbolicIOField "Campo ES simbólico_4" at 25,245 size 290x21
   TextField "Campo de texto_1" at 272,362 size 72x27
   Button "Botón_1" at 192,442 size 48x38
   Button "Botón_2" at 192,402 size 48x38
   TextField "Campo de texto_2" at 88,426 size 84x27
   GraphicIOField "Campo ES gráfico_1" at 300,402 size 16x78
   GraphicIOField "Campo ES gráfico_4" at 380,402 size 16x78
   TextField "Campo de texto_10" at 368,363 size 40x27
   SymbolicIOField "Campo ES simbólico_1" at 15,290 size 424x37
   Button "Botón_3" at 396,106 size 40x38
   Button "Botón_4" at 306,600 size 96x35
   TextField "Campo de texto_6" at 32,510 size 326x27
   TextField "Campo de texto_3" at 32,343 size 158x27
   TextField "Campo de texto_16" at 521,10 size 279x27
   Button "Botón_5" at 306,665 size 96x35
   TextField "Campo de texto_4" at 32,570 size 231x27
   TextField "Campo de texto_5" at 32,635 size 231x27
   IOField "Campo ES_7" at 20,535 size 173x35
   IOField "Campo ES_1" at 200,535 size 80x35
   IOField "Campo ES_2" at 20,595 size 173x35
   IOField "Campo ES_3" at 20,660 size 173x35

screen "MTA-ALTAMC002" 1280x800, template "Plantilla-Alta-Cmp"
   TextField "Campo de texto_1" at 266,362 size 72x27
   TextField "Campo de texto_2" at 82,426 size 84x27
   TextField "Campo de texto_10" at 362,363 size 40x27
   TextField "Campo de texto_6" at 32,510 size 326x27
   TextField "Campo de texto_3" at 26,343 size 158x27
   Button "Botón_1" at 186,442 size 48x38
   Button "Botón_2" at 186,402 size 48x38
   Button "Botón_3" at 390,106 size 40x38
   Button "Botón_4" at 306,600 size 96x35
   GraphicIOField "Campo ES gráfico_1" at 294,402 size 16x78
   GraphicIOField "Campo ES gráfico_4" at 374,402 size 16x78
   SymbolicIOField "Campo ES simbólico_1" at 9,290 size 424x37
   TextField "Campo de texto_16" at 521,10 size 279x27
   TextField "Campo de texto_4" at 32,570 size 231x27
   TextField "Campo de texto_5" at 32,635 size 231x27
   Button "Botón_5" at 306,665 size 96x35
   GraphicIOField "Campo ES gráfico_2" at 10,279 size 422x6
   SymbolicIOField "Campo ES simbólico_4" at 19,245 size 290x21
   Button "Botón_6" at 21,153 size 88x62
   Switch "Interruptor_1" at 150,166 size 37x37
   ScreenModuleView "Faceplate_6_1" at 342,235 size 76x34
   ScreenModuleView "Faceplate_7_1" at 213,157 size 208x70
   IOField "Campo ES_7" at 20,535 size 173x35
   IOField "Campo ES_1" at 200,535 size 80x35
   IOField "Campo ES_2" at 20,595 size 173x35
   IOField "Campo ES_3" at 20,660 size 173x35

screen "MTA-ALTAMC003" 1280x800, template "Plantilla-Alta-Cmp"
   Switch "Interruptor_1" at 150,119 size 37x37
   Button "Botón_6" at 13,106 size 88x62
   ScreenModuleView "Faceplate_6_1" at 342,236 size 76x34
   Button "Botón_1" at 186,441 size 48x38
   Button "Botón_2" at 186,401 size 48x38
   TextField "Campo de texto_6" at 266,362 size 72x27
   TextField "Campo de texto_7" at 82,426 size 84x27
   TextField "Campo de texto_8" at 362,363 size 40x27
   TextField "Campo de texto_9" at 32,510 size 326x27
   TextField "Campo de texto_11" at 26,343 size 158x27
   Button "Botón_7" at 390,58 size 40x38
   Button "Botón_8" at 306,600 size 96x35
   GraphicIOField "Campo ES gráfico_3" at 294,402 size 16x78
   GraphicIOField "Campo ES gráfico_5" at 374,402 size 16x78
   SymbolicIOField "Campo ES simbólico_2" at 9,290 size 424x37
   TextField "Campo de texto_16" at 521,10 size 270x27
   IOField "Campo ES_2" at 663,535 size 88x23
   TextField "Campo de texto_1" at 504,520 size 143x50
   Button "Botón_3" at 306,665 size 96x35
   TextField "Campo de texto_4" at 32,570 size 231x27
   TextField "Campo de texto_5" at 32,635 size 231x27
   GraphicIOField "Campo ES gráfico_2" at 10,280 size 422x6
   SymbolicIOField "Campo ES simbólico_4" at 19,246 size 290x21
   IOField "Campo ES_7" at 20,535 size 173x35
   IOField "Campo ES_1" at 200,535 size 80x35
   IOField "Campo ES_3" at 20,595 size 173x35
   IOField "Campo ES_4" at 20,660 size 173x35
   Switch "Interruptor_2" at 19,168 size 160x36
   ScreenModuleView "Faceplate_10_1" at 206,110 size 209x118

screen "MTA-ALTAMC004" 1280x800, template "Plantilla-Alta-Cmp"
   Button "Botón_1" at 186,441 size 48x38
   Button "Botón_2" at 186,401 size 48x38
   Button "Botón_7" at 390,106 size 40x38
   Button "Botón_8" at 300,600 size 96x35
   TextField "Campo de texto_6" at 266,362 size 72x27
   TextField "Campo de texto_7" at 82,426 size 84x27
   TextField "Campo de texto_8" at 362,363 size 40x27
   TextField "Campo de texto_11" at 26,343 size 158x27
   GraphicIOField "Campo ES gráfico_3" at 294,402 size 16x78
   GraphicIOField "Campo ES gráfico_5" at 374,402 size 16x78
   SymbolicIOField "Campo ES simbólico_2" at 9,290 size 424x37
   TextField "Campo de texto_16" at 521,10 size 279x27
   TextField "Campo de texto_1" at 32,510 size 326x27
   TextField "Campo de texto_4" at 32,570 size 231x27
   TextField "Campo de texto_5" at 32,635 size 231x27
   Button "Botón_3" at 300,665 size 96x35
   GraphicIOField "Campo ES gráfico_2" at 10,280 size 422x6
   SymbolicIOField "Campo ES simbólico_4" at 19,246 size 290x21
   Button "Botón_6" at 13,154 size 88x62
   Switch "Interruptor_1" at 150,167 size 37x37
   ScreenModuleView "Faceplate_6_1" at 342,236 size 76x34
   ScreenModuleView "Faceplate_7_1" at 213,158 size 208x70
   IOField "Campo ES_7" at 20,535 size 173x35
   IOField "Campo ES_1" at 200,535 size 80x35
   IOField "Campo ES_2" at 20,595 size 173x35
   IOField "Campo ES_3" at 20,660 size 173x35

screen "MTA-ALTAMC005" 1280x800, template "Plantilla-Alta-Cmp"
   Button "Botón_1" at 186,441 size 48x38
   Button "Botón_2" at 186,401 size 48x38
   Button "Botón_7" at 390,106 size 40x38
   Button "Botón_8" at 310,600 size 96x35
   TextField "Campo de texto_6" at 266,362 size 72x27
   TextField "Campo de texto_7" at 82,426 size 84x27
   TextField "Campo de texto_8" at 362,363 size 40x27
   TextField "Campo de texto_11" at 26,343 size 158x27
   GraphicIOField "Campo ES gráfico_3" at 294,402 size 16x78
   GraphicIOField "Campo ES gráfico_5" at 374,402 size 16x78
   SymbolicIOField "Campo ES simbólico_2" at 9,290 size 424x37
   TextField "Campo de texto_16" at 521,10 size 279x27
   TextField "Campo de texto_1" at 36,510 size 326x27
   TextField "Campo de texto_4" at 36,570 size 231x27
   TextField "Campo de texto_5" at 36,635 size 231x27
   Button "Botón_3" at 310,665 size 96x35
   GraphicIOField "Campo ES gráfico_2" at 10,280 size 422x6
   SymbolicIOField "Campo ES simbólico_4" at 19,246 size 290x21
   Button "Botón_6" at 13,154 size 88x62
   Switch "Interruptor_1" at 150,167 size 37x37
   ScreenModuleView "Faceplate_6_1" at 342,236 size 76x34
   ScreenModuleView "Faceplate_7_1" at 213,158 size 207x70
   IOField "Campo ES_7" at 24,535 size 173x35
   IOField "Campo ES_1" at 204,535 size 80x35
   IOField "Campo ES_2" at 24,595 size 173x35
   IOField "Campo ES_3" at 24,660 size 173x35

screen "MTA-Avisos" 1280x800, template "Plantilla"
   AlarmView "Visor de avisos_1" at 61,61 size 1174x631
   TextField "Campo de texto_16" at 613,9 size 54x27

screen "MTA-Avisos-Histórico" 1280x800, template "Plantilla"
   AlarmView "Visor de avisos_1" at 61,61 size 1174x631
   TextField "Campo de texto_16" at 573,9 size 157x27

screen "MTA-AyudaCFG1" 1280x800, template "Plantilla"
   TextField "Campo de texto_1" at 66,128 size 540x220
   TextField "Campo de texto_2" at 42,112 size 507x27
   TextField "Campo de texto_3" at 66,416 size 508x220
   TextField "Campo de texto_4" at 42,400 size 235x27
   TextField "Campo de texto_5" at 905,92 size 123x32
   TextField "Campo de texto_6" at 905,172 size 123x32
   TextField "Campo de texto_7" at 905,252 size 123x32
   TextField "Campo de texto_8" at 905,332 size 123x32
   TextField "Campo de texto_9" at 905,412 size 123x32
   TextField "Campo de texto_11" at 1148,498 size 88x32
   TextField "Campo de texto_12" at 708,557 size 128x18
   TextField "Campo de texto_13" at 708,611 size 122x18
   TextField "Campo de texto_14" at 1162,199 size 85x46
   TextField "Campo de texto_15" at 658,199 size 140x46
   Button "Botón_12" at 1089,638 size 160x49
   TextField "Campo de texto_16" at 414,9 size 455x27
   TextField "Campo de texto_10" at 905,492 size 123x32

screen "MTA-AyudaCmpAlta" 1280x800, template "Plantilla"
   Switch "Interruptor_1" at 1192,363 size 40x40
   GraphicIOField "Campo ES gráfico_6" at 763,381 size 9x45
   GraphicIOField "Campo ES gráfico_9" at 772,381 size 9x45
   GraphicView "Visor de gráficos_1" at 660,384 size 28x27
   TextField "Campo de texto_6" at 285,315 size 125x61
   TextField "Campo de texto_10" at 413,297 size 113x61
   TextField "Campo de texto_1" at 532,218 size 108x80
   GraphicView "Visor de gráficos_3" at 694,382 size 28x30
   GraphicView "Visor de gráficos_4" at 726,382 size 28x30
   GraphicView "Visor de gráficos_5" at 126,91 size 28x30
   GraphicView "Visor de gráficos_7" at 94,91 size 28x30
   GraphicView "Visor de gráficos_8" at 126,131 size 28x30
   GraphicView "Visor de gráficos_9" at 94,131 size 28x30
   GraphicView "Visor de gráficos_10" at 126,171 size 28x30
   GraphicView "Visor de gráficos_11" at 94,171 size 28x30
   GraphicView "Visor de gráficos_12" at 126,211 size 28x30
   GraphicView "Visor de gráficos_13" at 94,211 size 28x30
   GraphicView "Visor de gráficos_14" at 126,171 size 28x30
   GraphicIOField "Plantilla_Campo ES gráfico_5" at 897,433 size 65x60
   GraphicView "Visor de gráficos_2" at 924,363 size 260x142
   GraphicView "Visor de gráficos_6" at 971,83 size 262x142
   TextField "Campo de texto_7" at 607,463 size 54x42
   TextField "Campo de texto_11" at 1067,286 size 199x76
   TextField "Campo de texto_12" at 1056,264 size 210x42
   TextField "Campo de texto_13" at 695,98 size 210x42
   TextField "Campo de texto_16" at 926,529 size 134x42
   TextField "Campo de texto_18" at 529,9 size 241x27
   TextField "Campo de texto_3" at 703,239 size 90x80
   TextField "Campo de texto_4" at 815,215 size 95x80
   TextField "Campo de texto_5" at 700,485 size 129x61
   TextField "Campo de texto_2" at 223,92 size 170x42
   TextField "Campo de texto_8" at 223,132 size 284x42
   TextField "Campo de texto_9" at 223,172 size 268x42
   TextField "Campo de texto_14" at 223,212 size 122x42
   TextField "Campo de texto_15" at 561,383 size 61x22
   Button "Botón_3" at 95,559 size 280x70
   GraphicIOField "Campo ES gráfico_4" at 421,438 size 374x6
   SymbolicIOField "Campo ES simbólico_4" at 440,410 size 178x21
   TextField "Campo de texto_19" at 434,377 size 66x32
   IOField "Campo ES_6" at 662,413 size 85x19

screen "MTA-AyudaCmpAlta_1" 1280x800, template "Plantilla"
   TextField "Campo de texto_18" at 529,9 size 241x27
   TextField "Campo de texto_5" at 466,549 size 701x99
   TextField "Campo de texto_1" at 286,362 size 72x27
   TextField "Campo de texto_2" at 102,426 size 84x27
   TextField "Campo de texto_10" at 382,363 size 40x27
   TextField "Campo de texto_6" at 46,520 size 326x27
   TextField "Campo de texto_3" at 46,343 size 158x27
   Button "Botón_1" at 206,442 size 48x38
   Button "Botón_2" at 206,402 size 48x38
   Button "Botón_3" at 410,106 size 40x38
   Button "Botón_4" at 320,558 size 96x70
   GraphicIOField "Campo ES gráfico_1" at 314,402 size 16x78
   GraphicIOField "Campo ES gráfico_2" at 394,402 size 16x78
   TextField "Campo de texto_4" at 466,381 size 709x80
   TextField "Campo de texto_7" at 466,150 size 658x61
   TextField "Campo de texto_8" at 466,222 size 812x99
   TextField "Campo de texto_9" at 202,296 size 76x27
   GraphicIOField "Campo ES gráfico_3" at 30,279 size 422x6
   SymbolicIOField "Campo ES simbólico_2" at 39,245 size 290x21
   Button "Botón_6" at 41,153 size 88x62
   Switch "Interruptor_1" at 170,166 size 37x37
   ScreenModuleView "Faceplate_7_1" at 241,157 size 200x70
   IOField "Campo ES_7" at 88,558 size 173x35
   IOField "Campo ES_1" at 103,590 size 173x35
   GraphicView "Visor de gráficos_12" at 356,232 size 36x38
   GraphicView "Visor de gráficos_13" at 396,232 size 36x38

screen "MTA-AyudaColores" 1280x800, template "Plantilla"
   GraphicView "Visor de gráficos_1" at 156,507 size 64x58
   GraphicView "Visor de gráficos_3" at 156,251 size 64x58
   GraphicView "Visor de gráficos_4" at 156,315 size 64x58
   GraphicView "Visor de gráficos_5" at 156,187 size 64x58
   GraphicView "Visor de gráficos_6" at 156,379 size 64x58
   GraphicView "Visor de gráficos_7" at 156,443 size 64x58
   TextField "Campo de texto_1" at 234,518 size 172x42
   TextField "Campo de texto_2" at 130,112 size 233x32
   TextField "Campo de texto_3" at 234,262 size 75x42
   TextField "Campo de texto_4" at 234,326 size 431x42
   TextField "Campo de texto_5" at 234,198 size 99x42
   TextField "Campo de texto_6" at 234,390 size 56x42
   TextField "Campo de texto_7" at 234,454 size 77x42
   TextField "Campo de texto_8" at 130,598 size 666x58
   TextField "Campo de texto_9" at 130,646 size 1002x40
   TextField "Campo de texto_16" at 542,9 size 200x27

screen "MTA-AyudaMotores" 1280x800, template "Plantilla"
   TextField "Campo de texto_5" at 159,478 size 343x42
   TextField "Campo de texto_8" at 50,294 size 461x58
   TextField "Campo de texto_9" at 882,291 size 279x58
   GraphicView "Visor de gráficos_2" at 624,407 size 64x103
   GraphicIOField "Plantilla_Campo ES gráfico_4" at 660,481 size 81x68
   SymbolicIOField "Campo ES simbólico_3" at 572,220 size 220x29
   TextField "Campo de texto_10" at 575,161 size 52x23
   TextField "Campo de texto_17" at 573,193 size 146x18
   ScreenModuleView "ControlMotor-NoAUTO_4" at 599,262 size 171x108
   TextField "Campo de texto_1" at 39,261 size 436x42
   TextField "Campo de texto_2" at 871,261 size 179x42
   TextField "Campo de texto_3" at 871,373 size 160x42
   TextField "Campo de texto_4" at 119,205 size 376x42
   TextField "Campo de texto_6" at 871,165 size 251x23
   TextField "Campo de texto_7" at 871,197 size 135x42
   TextField "Campo de texto_16" at 573,9 size 135x27